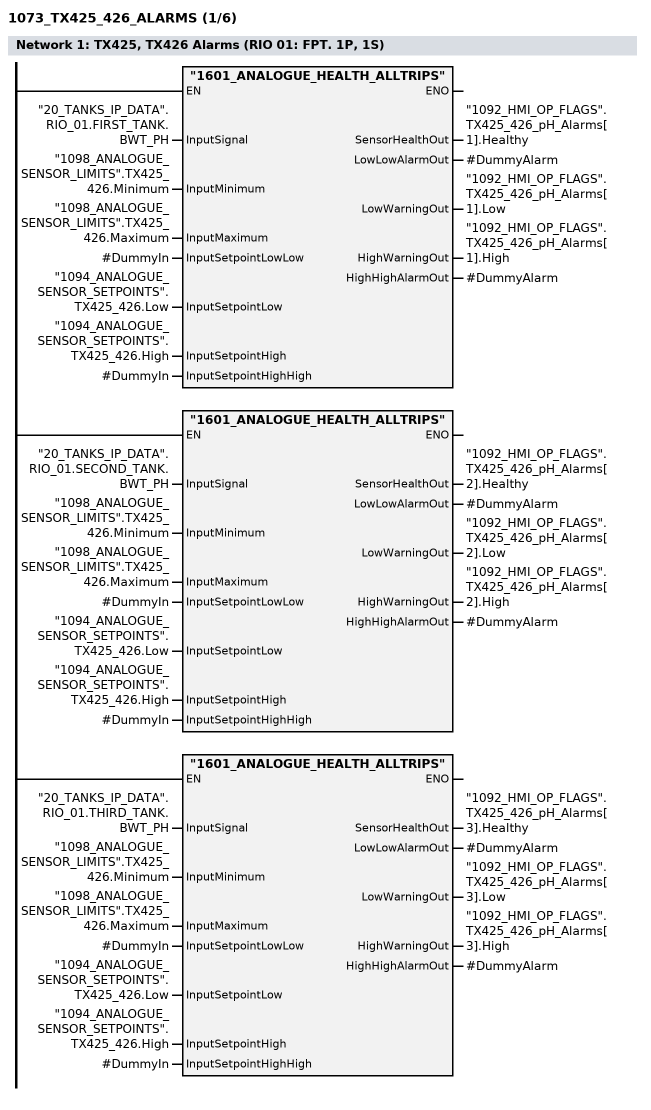
   RUNG wire#powerrail
      "1601_ANALOGUE_HEALTH_ALLTRIPS"(InputSignal := "20_TANKS_IP_DATA".RIO_01.FIRST_TANK.BWT_PH, InputMinimum := "1098_ANALOGUE_SENSOR_LIMITS".TX425_426.Minimum, InputMaximum := "1098_ANALOGUE_SENSOR_LIMITS".TX425_426.Maximum, InputSetpointLowLow := #DummyIn, InputSetpointLow := "1094_ANALOGUE_SENSOR_SETPOINTS".TX425_426.Low, InputSetpointHigh := "1094_ANALOGUE_SENSOR_SETPOINTS".TX425_426.High, InputSetpointHighHigh := #DummyIn, SensorHealthOut => "1092_HMI_OP_FLAGS".TX425_426_pH_Alarms[1].Healthy, LowLowAlarmOut => #DummyAlarm, LowWarningOut => "1092_HMI_OP_FLAGS".TX425_426_pH_Alarms[1].Low, HighWarningOut => "1092_HMI_OP_FLAGS".TX425_426_pH_Alarms[1].High, HighHighAlarmOut => #DummyAlarm)
   END_RUNG
   RUNG wire#powerrail
      "1601_ANALOGUE_HEALTH_ALLTRIPS"(InputSignal := "20_TANKS_IP_DATA".RIO_01.SECOND_TANK.BWT_PH, InputMinimum := "1098_ANALOGUE_SENSOR_LIMITS".TX425_426.Minimum, InputMaximum := "1098_ANALOGUE_SENSOR_LIMITS".TX425_426.Maximum, InputSetpointLowLow := #DummyIn, InputSetpointLow := "1094_ANALOGUE_SENSOR_SETPOINTS".TX425_426.Low, InputSetpointHigh := "1094_ANALOGUE_SENSOR_SETPOINTS".TX425_426.High, InputSetpointHighHigh := #DummyIn, SensorHealthOut => "1092_HMI_OP_FLAGS".TX425_426_pH_Alarms[2].Healthy, LowLowAlarmOut => #DummyAlarm, LowWarningOut => "1092_HMI_OP_FLAGS".TX425_426_pH_Alarms[2].Low, HighWarningOut => "1092_HMI_OP_FLAGS".TX425_426_pH_Alarms[2].High, HighHighAlarmOut => #DummyAlarm)
   END_RUNG
   RUNG wire#powerrail
      "1601_ANALOGUE_HEALTH_ALLTRIPS"(InputSignal := "20_TANKS_IP_DATA".RIO_01.THIRD_TANK.BWT_PH, InputMinimum := "1098_ANALOGUE_SENSOR_LIMITS".TX425_426.Minimum, InputMaximum := "1098_ANALOGUE_SENSOR_LIMITS".TX425_426.Maximum, InputSetpointLowLow := #DummyIn, InputSetpointLow := "1094_ANALOGUE_SENSOR_SETPOINTS".TX425_426.Low, InputSetpointHigh := "1094_ANALOGUE_SENSOR_SETPOINTS".TX425_426.High, InputSetpointHighHigh := #DummyIn, SensorHealthOut => "1092_HMI_OP_FLAGS".TX425_426_pH_Alarms[3].Healthy, LowLowAlarmOut => #DummyAlarm, LowWarningOut => "1092_HMI_OP_FLAGS".TX425_426_pH_Alarms[3].Low, HighWarningOut => "1092_HMI_OP_FLAGS".TX425_426_pH_Alarms[3].High, HighHighAlarmOut => #DummyAlarm)
   END_RUNG
   // the same network as SCL:
   "1601_ANALOGUE_HEALTH_ALLTRIPS"(InputSignal := "20_TANKS_IP_DATA".RIO_01.FIRST_TANK.BWT_PH,
                           InputMinimum := "1098_ANALOGUE_SENSOR_LIMITS".TX425_426.Minimum,
                           InputMaximum := "1098_ANALOGUE_SENSOR_LIMITS".TX425_426.Maximum,
                           InputSetpointLowLow := #DummyIn,
                           InputSetpointLow := "1094_ANALOGUE_SENSOR_SETPOINTS".TX425_426.Low,
                           InputSetpointHigh := "1094_ANALOGUE_SENSOR_SETPOINTS".TX425_426.High,
                           InputSetpointHighHigh := #DummyIn,
                           SensorHealthOut => "1092_HMI_OP_FLAGS".TX425_426_pH_Alarms[1].Healthy,
                           LowLowAlarmOut => #DummyAlarm,
                           LowWarningOut => "1092_HMI_OP_FLAGS".TX425_426_pH_Alarms[1].Low,
                           HighWarningOut => "1092_HMI_OP_FLAGS".TX425_426_pH_Alarms[1].High,
                           HighHighAlarmOut => #DummyAlarm);
   "1601_ANALOGUE_HEALTH_ALLTRIPS"(InputSignal := "20_TANKS_IP_DATA".RIO_01.SECOND_TANK.BWT_PH,
                           InputMinimum := "1098_ANALOGUE_SENSOR_LIMITS".TX425_426.Minimum,
                           InputMaximum := "1098_ANALOGUE_SENSOR_LIMITS".TX425_426.Maximum,
                           InputSetpointLowLow := #DummyIn,
                           InputSetpointLow := "1094_ANALOGUE_SENSOR_SETPOINTS".TX425_426.Low,
                           InputSetpointHigh := "1094_ANALOGUE_SENSOR_SETPOINTS".TX425_426.High,
                           InputSetpointHighHigh := #DummyIn,
                           SensorHealthOut => "1092_HMI_OP_FLAGS".TX425_426_pH_Alarms[2].Healthy,
                           LowLowAlarmOut => #DummyAlarm,
                           LowWarningOut => "1092_HMI_OP_FLAGS".TX425_426_pH_Alarms[2].Low,
                           HighWarningOut => "1092_HMI_OP_FLAGS".TX425_426_pH_Alarms[2].High,
                           HighHighAlarmOut => #DummyAlarm);
   "1601_ANALOGUE_HEALTH_ALLTRIPS"(InputSignal := "20_TANKS_IP_DATA".RIO_01.THIRD_TANK.BWT_PH,
                           InputMinimum := "1098_ANALOGUE_SENSOR_LIMITS".TX425_426.Minimum,
                           InputMaximum := "1098_ANALOGUE_SENSOR_LIMITS".TX425_426.Maximum,
                           InputSetpointLowLow := #DummyIn,
                           InputSetpointLow := "1094_ANALOGUE_SENSOR_SETPOINTS".TX425_426.Low,
                           InputSetpointHigh := "1094_ANALOGUE_SENSOR_SETPOINTS".TX425_426.High,
                           InputSetpointHighHigh := #DummyIn,
                           SensorHealthOut => "1092_HMI_OP_FLAGS".TX425_426_pH_Alarms[3].Healthy,
                           LowLowAlarmOut => #DummyAlarm,
                           LowWarningOut => "1092_HMI_OP_FLAGS".TX425_426_pH_Alarms[3].Low,
                           HighWarningOut => "1092_HMI_OP_FLAGS".TX425_426_pH_Alarms[3].High,
                           HighHighAlarmOut => #DummyAlarm);
END_REGION

REGION Network 2: TX425, TX426 Alarms (RIO 02: 2P, 2S)
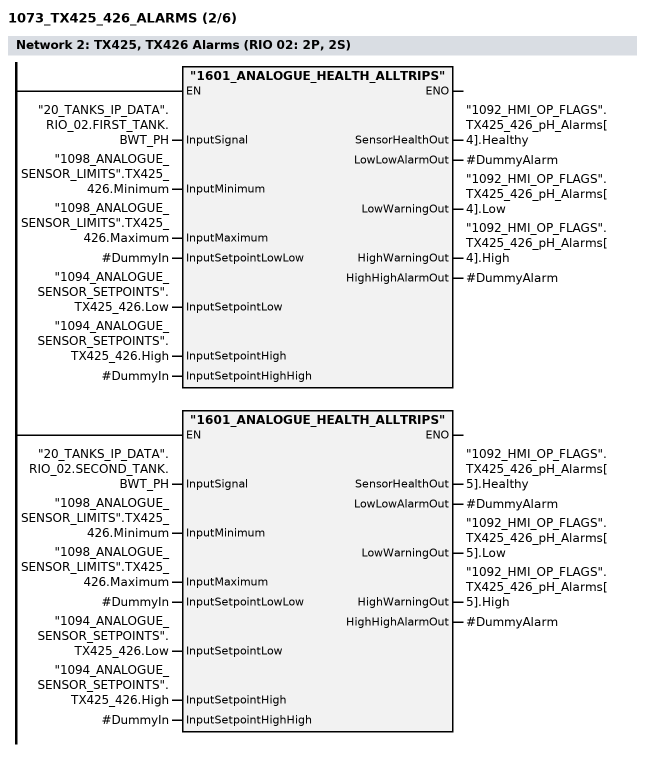
   RUNG wire#powerrail
      "1601_ANALOGUE_HEALTH_ALLTRIPS"(InputSignal := "20_TANKS_IP_DATA".RIO_02.FIRST_TANK.BWT_PH, InputMinimum := "1098_ANALOGUE_SENSOR_LIMITS".TX425_426.Minimum, InputMaximum := "1098_ANALOGUE_SENSOR_LIMITS".TX425_426.Maximum, InputSetpointLowLow := #DummyIn, InputSetpointLow := "1094_ANALOGUE_SENSOR_SETPOINTS".TX425_426.Low, InputSetpointHigh := "1094_ANALOGUE_SENSOR_SETPOINTS".TX425_426.High, InputSetpointHighHigh := #DummyIn, SensorHealthOut => "1092_HMI_OP_FLAGS".TX425_426_pH_Alarms[4].Healthy, LowLowAlarmOut => #DummyAlarm, LowWarningOut => "1092_HMI_OP_FLAGS".TX425_426_pH_Alarms[4].Low, HighWarningOut => "1092_HMI_OP_FLAGS".TX425_426_pH_Alarms[4].High, HighHighAlarmOut => #DummyAlarm)
   END_RUNG
   RUNG wire#powerrail
      "1601_ANALOGUE_HEALTH_ALLTRIPS"(InputSignal := "20_TANKS_IP_DATA".RIO_02.SECOND_TANK.BWT_PH, InputMinimum := "1098_ANALOGUE_SENSOR_LIMITS".TX425_426.Minimum, InputMaximum := "1098_ANALOGUE_SENSOR_LIMITS".TX425_426.Maximum, InputSetpointLowLow := #DummyIn, InputSetpointLow := "1094_ANALOGUE_SENSOR_SETPOINTS".TX425_426.Low, InputSetpointHigh := "1094_ANALOGUE_SENSOR_SETPOINTS".TX425_426.High, InputSetpointHighHigh := #DummyIn, SensorHealthOut => "1092_HMI_OP_FLAGS".TX425_426_pH_Alarms[5].Healthy, LowLowAlarmOut => #DummyAlarm, LowWarningOut => "1092_HMI_OP_FLAGS".TX425_426_pH_Alarms[5].Low, HighWarningOut => "1092_HMI_OP_FLAGS".TX425_426_pH_Alarms[5].High, HighHighAlarmOut => #DummyAlarm)
   END_RUNG
   // the same network as SCL:
   "1601_ANALOGUE_HEALTH_ALLTRIPS"(InputSignal := "20_TANKS_IP_DATA".RIO_02.FIRST_TANK.BWT_PH,
                           InputMinimum := "1098_ANALOGUE_SENSOR_LIMITS".TX425_426.Minimum,
                           InputMaximum := "1098_ANALOGUE_SENSOR_LIMITS".TX425_426.Maximum,
                           InputSetpointLowLow := #DummyIn,
                           InputSetpointLow := "1094_ANALOGUE_SENSOR_SETPOINTS".TX425_426.Low,
                           InputSetpointHigh := "1094_ANALOGUE_SENSOR_SETPOINTS".TX425_426.High,
                           InputSetpointHighHigh := #DummyIn,
                           SensorHealthOut => "1092_HMI_OP_FLAGS".TX425_426_pH_Alarms[4].Healthy,
                           LowLowAlarmOut => #DummyAlarm,
                           LowWarningOut => "1092_HMI_OP_FLAGS".TX425_426_pH_Alarms[4].Low,
                           HighWarningOut => "1092_HMI_OP_FLAGS".TX425_426_pH_Alarms[4].High,
                           HighHighAlarmOut => #DummyAlarm);
   "1601_ANALOGUE_HEALTH_ALLTRIPS"(InputSignal := "20_TANKS_IP_DATA".RIO_02.SECOND_TANK.BWT_PH,
                           InputMinimum := "1098_ANALOGUE_SENSOR_LIMITS".TX425_426.Minimum,
                           InputMaximum := "1098_ANALOGUE_SENSOR_LIMITS".TX425_426.Maximum,
                           InputSetpointLowLow := #DummyIn,
                           InputSetpointLow := "1094_ANALOGUE_SENSOR_SETPOINTS".TX425_426.Low,
                           InputSetpointHigh := "1094_ANALOGUE_SENSOR_SETPOINTS".TX425_426.High,
                           InputSetpointHighHigh := #DummyIn,
                           SensorHealthOut => "1092_HMI_OP_FLAGS".TX425_426_pH_Alarms[5].Healthy,
                           LowLowAlarmOut => #DummyAlarm,
                           LowWarningOut => "1092_HMI_OP_FLAGS".TX425_426_pH_Alarms[5].Low,
                           HighWarningOut => "1092_HMI_OP_FLAGS".TX425_426_pH_Alarms[5].High,
                           HighHighAlarmOut => #DummyAlarm);
END_REGION

REGION Network 3: TX425, TX426 Alarms (RIO 03: 3P, 3S)
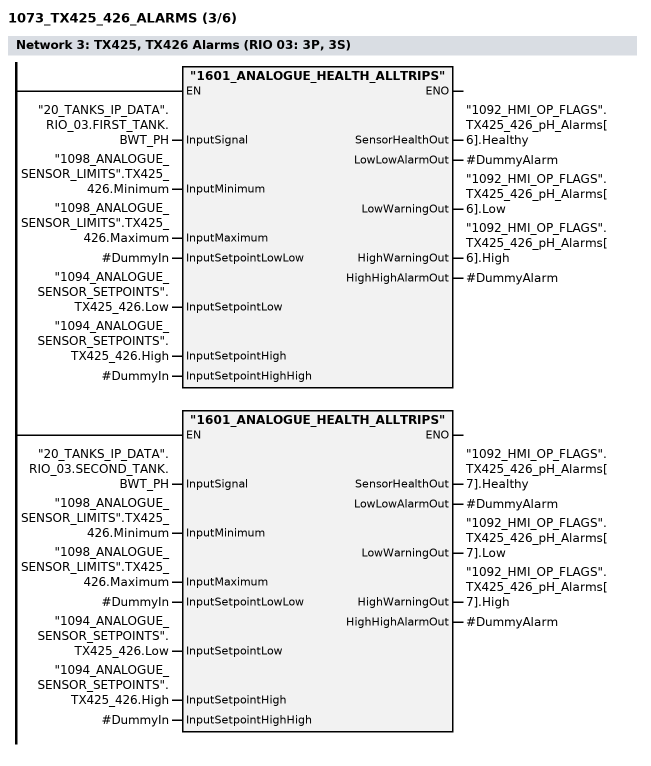
   RUNG wire#powerrail
      "1601_ANALOGUE_HEALTH_ALLTRIPS"(InputSignal := "20_TANKS_IP_DATA".RIO_03.FIRST_TANK.BWT_PH, InputMinimum := "1098_ANALOGUE_SENSOR_LIMITS".TX425_426.Minimum, InputMaximum := "1098_ANALOGUE_SENSOR_LIMITS".TX425_426.Maximum, InputSetpointLowLow := #DummyIn, InputSetpointLow := "1094_ANALOGUE_SENSOR_SETPOINTS".TX425_426.Low, InputSetpointHigh := "1094_ANALOGUE_SENSOR_SETPOINTS".TX425_426.High, InputSetpointHighHigh := #DummyIn, SensorHealthOut => "1092_HMI_OP_FLAGS".TX425_426_pH_Alarms[6].Healthy, LowLowAlarmOut => #DummyAlarm, LowWarningOut => "1092_HMI_OP_FLAGS".TX425_426_pH_Alarms[6].Low, HighWarningOut => "1092_HMI_OP_FLAGS".TX425_426_pH_Alarms[6].High, HighHighAlarmOut => #DummyAlarm)
   END_RUNG
   RUNG wire#powerrail
      "1601_ANALOGUE_HEALTH_ALLTRIPS"(InputSignal := "20_TANKS_IP_DATA".RIO_03.SECOND_TANK.BWT_PH, InputMinimum := "1098_ANALOGUE_SENSOR_LIMITS".TX425_426.Minimum, InputMaximum := "1098_ANALOGUE_SENSOR_LIMITS".TX425_426.Maximum, InputSetpointLowLow := #DummyIn, InputSetpointLow := "1094_ANALOGUE_SENSOR_SETPOINTS".TX425_426.Low, InputSetpointHigh := "1094_ANALOGUE_SENSOR_SETPOINTS".TX425_426.High, InputSetpointHighHigh := #DummyIn, SensorHealthOut => "1092_HMI_OP_FLAGS".TX425_426_pH_Alarms[7].Healthy, LowLowAlarmOut => #DummyAlarm, LowWarningOut => "1092_HMI_OP_FLAGS".TX425_426_pH_Alarms[7].Low, HighWarningOut => "1092_HMI_OP_FLAGS".TX425_426_pH_Alarms[7].High, HighHighAlarmOut => #DummyAlarm)
   END_RUNG
   // the same network as SCL:
   "1601_ANALOGUE_HEALTH_ALLTRIPS"(InputSignal := "20_TANKS_IP_DATA".RIO_03.FIRST_TANK.BWT_PH,
                           InputMinimum := "1098_ANALOGUE_SENSOR_LIMITS".TX425_426.Minimum,
                           InputMaximum := "1098_ANALOGUE_SENSOR_LIMITS".TX425_426.Maximum,
                           InputSetpointLowLow := #DummyIn,
                           InputSetpointLow := "1094_ANALOGUE_SENSOR_SETPOINTS".TX425_426.Low,
                           InputSetpointHigh := "1094_ANALOGUE_SENSOR_SETPOINTS".TX425_426.High,
                           InputSetpointHighHigh := #DummyIn,
                           SensorHealthOut => "1092_HMI_OP_FLAGS".TX425_426_pH_Alarms[6].Healthy,
                           LowLowAlarmOut => #DummyAlarm,
                           LowWarningOut => "1092_HMI_OP_FLAGS".TX425_426_pH_Alarms[6].Low,
                           HighWarningOut => "1092_HMI_OP_FLAGS".TX425_426_pH_Alarms[6].High,
                           HighHighAlarmOut => #DummyAlarm);
   "1601_ANALOGUE_HEALTH_ALLTRIPS"(InputSignal := "20_TANKS_IP_DATA".RIO_03.SECOND_TANK.BWT_PH,
                           InputMinimum := "1098_ANALOGUE_SENSOR_LIMITS".TX425_426.Minimum,
                           InputMaximum := "1098_ANALOGUE_SENSOR_LIMITS".TX425_426.Maximum,
                           InputSetpointLowLow := #DummyIn,
                           InputSetpointLow := "1094_ANALOGUE_SENSOR_SETPOINTS".TX425_426.Low,
                           InputSetpointHigh := "1094_ANALOGUE_SENSOR_SETPOINTS".TX425_426.High,
                           InputSetpointHighHigh := #DummyIn,
                           SensorHealthOut => "1092_HMI_OP_FLAGS".TX425_426_pH_Alarms[7].Healthy,
                           LowLowAlarmOut => #DummyAlarm,
                           LowWarningOut => "1092_HMI_OP_FLAGS".TX425_426_pH_Alarms[7].Low,
                           HighWarningOut => "1092_HMI_OP_FLAGS".TX425_426_pH_Alarms[7].High,
                           HighHighAlarmOut => #DummyAlarm);
END_REGION

REGION Network 4: TX425, TX426 Alarms (RIO 04: 4P, 4S)
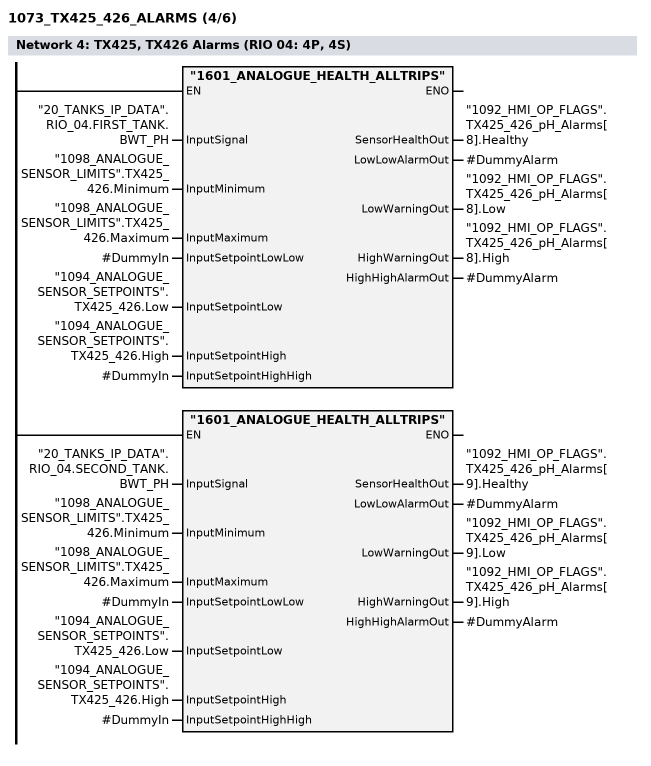
   RUNG wire#powerrail
      "1601_ANALOGUE_HEALTH_ALLTRIPS"(InputSignal := "20_TANKS_IP_DATA".RIO_04.FIRST_TANK.BWT_PH, InputMinimum := "1098_ANALOGUE_SENSOR_LIMITS".TX425_426.Minimum, InputMaximum := "1098_ANALOGUE_SENSOR_LIMITS".TX425_426.Maximum, InputSetpointLowLow := #DummyIn, InputSetpointLow := "1094_ANALOGUE_SENSOR_SETPOINTS".TX425_426.Low, InputSetpointHigh := "1094_ANALOGUE_SENSOR_SETPOINTS".TX425_426.High, InputSetpointHighHigh := #DummyIn, SensorHealthOut => "1092_HMI_OP_FLAGS".TX425_426_pH_Alarms[8].Healthy, LowLowAlarmOut => #DummyAlarm, LowWarningOut => "1092_HMI_OP_FLAGS".TX425_426_pH_Alarms[8].Low, HighWarningOut => "1092_HMI_OP_FLAGS".TX425_426_pH_Alarms[8].High, HighHighAlarmOut => #DummyAlarm)
   END_RUNG
   RUNG wire#powerrail
      "1601_ANALOGUE_HEALTH_ALLTRIPS"(InputSignal := "20_TANKS_IP_DATA".RIO_04.SECOND_TANK.BWT_PH, InputMinimum := "1098_ANALOGUE_SENSOR_LIMITS".TX425_426.Minimum, InputMaximum := "1098_ANALOGUE_SENSOR_LIMITS".TX425_426.Maximum, InputSetpointLowLow := #DummyIn, InputSetpointLow := "1094_ANALOGUE_SENSOR_SETPOINTS".TX425_426.Low, InputSetpointHigh := "1094_ANALOGUE_SENSOR_SETPOINTS".TX425_426.High, InputSetpointHighHigh := #DummyIn, SensorHealthOut => "1092_HMI_OP_FLAGS".TX425_426_pH_Alarms[9].Healthy, LowLowAlarmOut => #DummyAlarm, LowWarningOut => "1092_HMI_OP_FLAGS".TX425_426_pH_Alarms[9].Low, HighWarningOut => "1092_HMI_OP_FLAGS".TX425_426_pH_Alarms[9].High, HighHighAlarmOut => #DummyAlarm)
   END_RUNG
   // the same network as SCL:
   "1601_ANALOGUE_HEALTH_ALLTRIPS"(InputSignal := "20_TANKS_IP_DATA".RIO_04.FIRST_TANK.BWT_PH,
                           InputMinimum := "1098_ANALOGUE_SENSOR_LIMITS".TX425_426.Minimum,
                           InputMaximum := "1098_ANALOGUE_SENSOR_LIMITS".TX425_426.Maximum,
                           InputSetpointLowLow := #DummyIn,
                           InputSetpointLow := "1094_ANALOGUE_SENSOR_SETPOINTS".TX425_426.Low,
                           InputSetpointHigh := "1094_ANALOGUE_SENSOR_SETPOINTS".TX425_426.High,
                           InputSetpointHighHigh := #DummyIn,
                           SensorHealthOut => "1092_HMI_OP_FLAGS".TX425_426_pH_Alarms[8].Healthy,
                           LowLowAlarmOut => #DummyAlarm,
                           LowWarningOut => "1092_HMI_OP_FLAGS".TX425_426_pH_Alarms[8].Low,
                           HighWarningOut => "1092_HMI_OP_FLAGS".TX425_426_pH_Alarms[8].High,
                           HighHighAlarmOut => #DummyAlarm);
   "1601_ANALOGUE_HEALTH_ALLTRIPS"(InputSignal := "20_TANKS_IP_DATA".RIO_04.SECOND_TANK.BWT_PH,
                           InputMinimum := "1098_ANALOGUE_SENSOR_LIMITS".TX425_426.Minimum,
                           InputMaximum := "1098_ANALOGUE_SENSOR_LIMITS".TX425_426.Maximum,
                           InputSetpointLowLow := #DummyIn,
                           InputSetpointLow := "1094_ANALOGUE_SENSOR_SETPOINTS".TX425_426.Low,
                           InputSetpointHigh := "1094_ANALOGUE_SENSOR_SETPOINTS".TX425_426.High,
                           InputSetpointHighHigh := #DummyIn,
                           SensorHealthOut => "1092_HMI_OP_FLAGS".TX425_426_pH_Alarms[9].Healthy,
                           LowLowAlarmOut => #DummyAlarm,
                           LowWarningOut => "1092_HMI_OP_FLAGS".TX425_426_pH_Alarms[9].Low,
                           HighWarningOut => "1092_HMI_OP_FLAGS".TX425_426_pH_Alarms[9].High,
                           HighHighAlarmOut => #DummyAlarm);
END_REGION

REGION Network 5: TX425, TX426 Alarms (RIO 05: 5P, 5S)
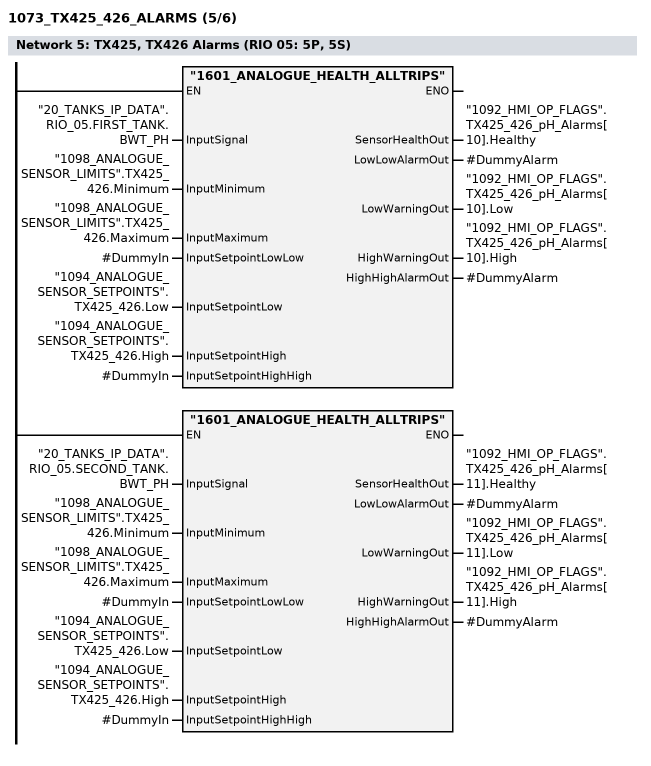
   RUNG wire#powerrail
      "1601_ANALOGUE_HEALTH_ALLTRIPS"(InputSignal := "20_TANKS_IP_DATA".RIO_05.FIRST_TANK.BWT_PH, InputMinimum := "1098_ANALOGUE_SENSOR_LIMITS".TX425_426.Minimum, InputMaximum := "1098_ANALOGUE_SENSOR_LIMITS".TX425_426.Maximum, InputSetpointLowLow := #DummyIn, InputSetpointLow := "1094_ANALOGUE_SENSOR_SETPOINTS".TX425_426.Low, InputSetpointHigh := "1094_ANALOGUE_SENSOR_SETPOINTS".TX425_426.High, InputSetpointHighHigh := #DummyIn, SensorHealthOut => "1092_HMI_OP_FLAGS".TX425_426_pH_Alarms[10].Healthy, LowLowAlarmOut => #DummyAlarm, LowWarningOut => "1092_HMI_OP_FLAGS".TX425_426_pH_Alarms[10].Low, HighWarningOut => "1092_HMI_OP_FLAGS".TX425_426_pH_Alarms[10].High, HighHighAlarmOut => #DummyAlarm)
   END_RUNG
   RUNG wire#powerrail
      "1601_ANALOGUE_HEALTH_ALLTRIPS"(InputSignal := "20_TANKS_IP_DATA".RIO_05.SECOND_TANK.BWT_PH, InputMinimum := "1098_ANALOGUE_SENSOR_LIMITS".TX425_426.Minimum, InputMaximum := "1098_ANALOGUE_SENSOR_LIMITS".TX425_426.Maximum, InputSetpointLowLow := #DummyIn, InputSetpointLow := "1094_ANALOGUE_SENSOR_SETPOINTS".TX425_426.Low, InputSetpointHigh := "1094_ANALOGUE_SENSOR_SETPOINTS".TX425_426.High, InputSetpointHighHigh := #DummyIn, SensorHealthOut => "1092_HMI_OP_FLAGS".TX425_426_pH_Alarms[11].Healthy, LowLowAlarmOut => #DummyAlarm, LowWarningOut => "1092_HMI_OP_FLAGS".TX425_426_pH_Alarms[11].Low, HighWarningOut => "1092_HMI_OP_FLAGS".TX425_426_pH_Alarms[11].High, HighHighAlarmOut => #DummyAlarm)
   END_RUNG
   // the same network as SCL:
   "1601_ANALOGUE_HEALTH_ALLTRIPS"(InputSignal := "20_TANKS_IP_DATA".RIO_05.FIRST_TANK.BWT_PH,
                           InputMinimum := "1098_ANALOGUE_SENSOR_LIMITS".TX425_426.Minimum,
                           InputMaximum := "1098_ANALOGUE_SENSOR_LIMITS".TX425_426.Maximum,
                           InputSetpointLowLow := #DummyIn,
                           InputSetpointLow := "1094_ANALOGUE_SENSOR_SETPOINTS".TX425_426.Low,
                           InputSetpointHigh := "1094_ANALOGUE_SENSOR_SETPOINTS".TX425_426.High,
                           InputSetpointHighHigh := #DummyIn,
                           SensorHealthOut => "1092_HMI_OP_FLAGS".TX425_426_pH_Alarms[10].Healthy,
                           LowLowAlarmOut => #DummyAlarm,
                           LowWarningOut => "1092_HMI_OP_FLAGS".TX425_426_pH_Alarms[10].Low,
                           HighWarningOut => "1092_HMI_OP_FLAGS".TX425_426_pH_Alarms[10].High,
                           HighHighAlarmOut => #DummyAlarm);
   "1601_ANALOGUE_HEALTH_ALLTRIPS"(InputSignal := "20_TANKS_IP_DATA".RIO_05.SECOND_TANK.BWT_PH,
                           InputMinimum := "1098_ANALOGUE_SENSOR_LIMITS".TX425_426.Minimum,
                           InputMaximum := "1098_ANALOGUE_SENSOR_LIMITS".TX425_426.Maximum,
                           InputSetpointLowLow := #DummyIn,
                           InputSetpointLow := "1094_ANALOGUE_SENSOR_SETPOINTS".TX425_426.Low,
                           InputSetpointHigh := "1094_ANALOGUE_SENSOR_SETPOINTS".TX425_426.High,
                           InputSetpointHighHigh := #DummyIn,
                           SensorHealthOut => "1092_HMI_OP_FLAGS".TX425_426_pH_Alarms[11].Healthy,
                           LowLowAlarmOut => #DummyAlarm,
                           LowWarningOut => "1092_HMI_OP_FLAGS".TX425_426_pH_Alarms[11].Low,
                           HighWarningOut => "1092_HMI_OP_FLAGS".TX425_426_pH_Alarms[11].High,
                           HighHighAlarmOut => #DummyAlarm);
END_REGION

REGION Network 6: TX425, TX426 Alarms (RIO 06: 6P, 6S)
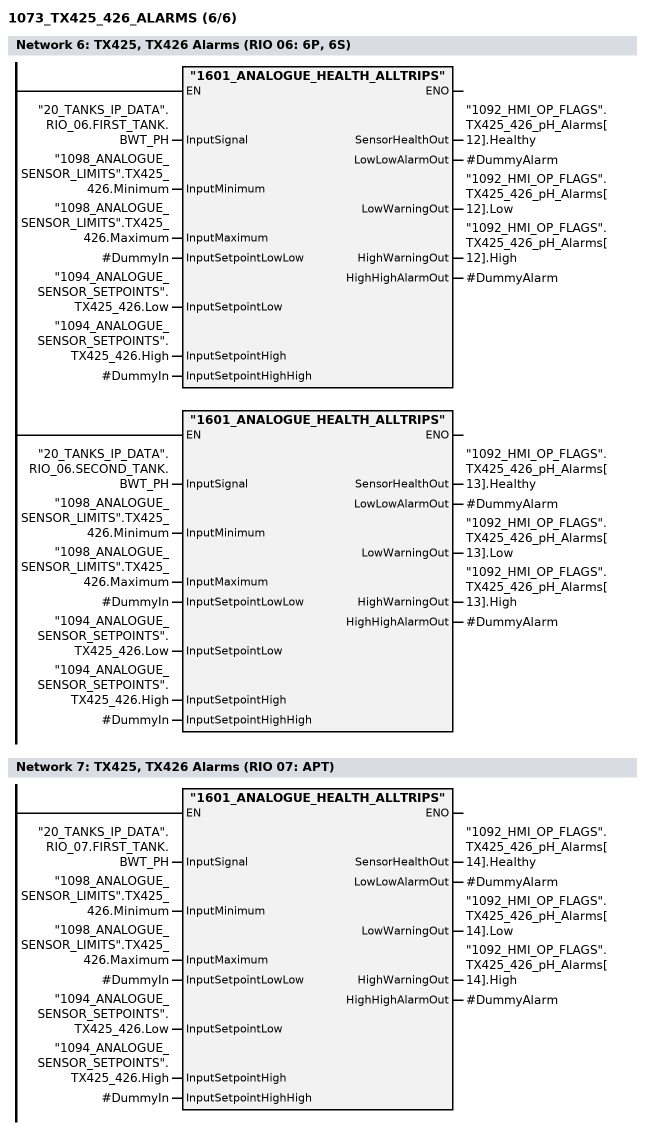
   RUNG wire#powerrail
      "1601_ANALOGUE_HEALTH_ALLTRIPS"(InputSignal := "20_TANKS_IP_DATA".RIO_06.FIRST_TANK.BWT_PH, InputMinimum := "1098_ANALOGUE_SENSOR_LIMITS".TX425_426.Minimum, InputMaximum := "1098_ANALOGUE_SENSOR_LIMITS".TX425_426.Maximum, InputSetpointLowLow := #DummyIn, InputSetpointLow := "1094_ANALOGUE_SENSOR_SETPOINTS".TX425_426.Low, InputSetpointHigh := "1094_ANALOGUE_SENSOR_SETPOINTS".TX425_426.High, InputSetpointHighHigh := #DummyIn, SensorHealthOut => "1092_HMI_OP_FLAGS".TX425_426_pH_Alarms[12].Healthy, LowLowAlarmOut => #DummyAlarm, LowWarningOut => "1092_HMI_OP_FLAGS".TX425_426_pH_Alarms[12].Low, HighWarningOut => "1092_HMI_OP_FLAGS".TX425_426_pH_Alarms[12].High, HighHighAlarmOut => #DummyAlarm)
   END_RUNG
   RUNG wire#powerrail
      "1601_ANALOGUE_HEALTH_ALLTRIPS"(InputSignal := "20_TANKS_IP_DATA".RIO_06.SECOND_TANK.BWT_PH, InputMinimum := "1098_ANALOGUE_SENSOR_LIMITS".TX425_426.Minimum, InputMaximum := "1098_ANALOGUE_SENSOR_LIMITS".TX425_426.Maximum, InputSetpointLowLow := #DummyIn, InputSetpointLow := "1094_ANALOGUE_SENSOR_SETPOINTS".TX425_426.Low, InputSetpointHigh := "1094_ANALOGUE_SENSOR_SETPOINTS".TX425_426.High, InputSetpointHighHigh := #DummyIn, SensorHealthOut => "1092_HMI_OP_FLAGS".TX425_426_pH_Alarms[13].Healthy, LowLowAlarmOut => #DummyAlarm, LowWarningOut => "1092_HMI_OP_FLAGS".TX425_426_pH_Alarms[13].Low, HighWarningOut => "1092_HMI_OP_FLAGS".TX425_426_pH_Alarms[13].High, HighHighAlarmOut => #DummyAlarm)
   END_RUNG
   // the same network as SCL:
   "1601_ANALOGUE_HEALTH_ALLTRIPS"(InputSignal := "20_TANKS_IP_DATA".RIO_06.FIRST_TANK.BWT_PH,
                           InputMinimum := "1098_ANALOGUE_SENSOR_LIMITS".TX425_426.Minimum,
                           InputMaximum := "1098_ANALOGUE_SENSOR_LIMITS".TX425_426.Maximum,
                           InputSetpointLowLow := #DummyIn,
                           InputSetpointLow := "1094_ANALOGUE_SENSOR_SETPOINTS".TX425_426.Low,
                           InputSetpointHigh := "1094_ANALOGUE_SENSOR_SETPOINTS".TX425_426.High,
                           InputSetpointHighHigh := #DummyIn,
                           SensorHealthOut => "1092_HMI_OP_FLAGS".TX425_426_pH_Alarms[12].Healthy,
                           LowLowAlarmOut => #DummyAlarm,
                           LowWarningOut => "1092_HMI_OP_FLAGS".TX425_426_pH_Alarms[12].Low,
                           HighWarningOut => "1092_HMI_OP_FLAGS".TX425_426_pH_Alarms[12].High,
                           HighHighAlarmOut => #DummyAlarm);
   "1601_ANALOGUE_HEALTH_ALLTRIPS"(InputSignal := "20_TANKS_IP_DATA".RIO_06.SECOND_TANK.BWT_PH,
                           InputMinimum := "1098_ANALOGUE_SENSOR_LIMITS".TX425_426.Minimum,
                           InputMaximum := "1098_ANALOGUE_SENSOR_LIMITS".TX425_426.Maximum,
                           InputSetpointLowLow := #DummyIn,
                           InputSetpointLow := "1094_ANALOGUE_SENSOR_SETPOINTS".TX425_426.Low,
                           InputSetpointHigh := "1094_ANALOGUE_SENSOR_SETPOINTS".TX425_426.High,
                           InputSetpointHighHigh := #DummyIn,
                           SensorHealthOut => "1092_HMI_OP_FLAGS".TX425_426_pH_Alarms[13].Healthy,
                           LowLowAlarmOut => #DummyAlarm,
                           LowWarningOut => "1092_HMI_OP_FLAGS".TX425_426_pH_Alarms[13].Low,
                           HighWarningOut => "1092_HMI_OP_FLAGS".TX425_426_pH_Alarms[13].High,
                           HighHighAlarmOut => #DummyAlarm);
END_REGION

REGION Network 7: TX425, TX426 Alarms (RIO 07: APT)
   RUNG wire#powerrail
      "1601_ANALOGUE_HEALTH_ALLTRIPS"(InputSignal := "20_TANKS_IP_DATA".RIO_07.FIRST_TANK.BWT_PH, InputMinimum := "1098_ANALOGUE_SENSOR_LIMITS".TX425_426.Minimum, InputMaximum := "1098_ANALOGUE_SENSOR_LIMITS".TX425_426.Maximum, InputSetpointLowLow := #DummyIn, InputSetpointLow := "1094_ANALOGUE_SENSOR_SETPOINTS".TX425_426.Low, InputSetpointHigh := "1094_ANALOGUE_SENSOR_SETPOINTS".TX425_426.High, InputSetpointHighHigh := #DummyIn, SensorHealthOut => "1092_HMI_OP_FLAGS".TX425_426_pH_Alarms[14].Healthy, LowLowAlarmOut => #DummyAlarm, LowWarningOut => "1092_HMI_OP_FLAGS".TX425_426_pH_Alarms[14].Low, HighWarningOut => "1092_HMI_OP_FLAGS".TX425_426_pH_Alarms[14].High, HighHighAlarmOut => #DummyAlarm)
   END_RUNG
   // the same network as SCL:
   "1601_ANALOGUE_HEALTH_ALLTRIPS"(InputSignal := "20_TANKS_IP_DATA".RIO_07.FIRST_TANK.BWT_PH,
                           InputMinimum := "1098_ANALOGUE_SENSOR_LIMITS".TX425_426.Minimum,
                           InputMaximum := "1098_ANALOGUE_SENSOR_LIMITS".TX425_426.Maximum,
                           InputSetpointLowLow := #DummyIn,
                           InputSetpointLow := "1094_ANALOGUE_SENSOR_SETPOINTS".TX425_426.Low,
                           InputSetpointHigh := "1094_ANALOGUE_SENSOR_SETPOINTS".TX425_426.High,
                           InputSetpointHighHigh := #DummyIn,
                           SensorHealthOut => "1092_HMI_OP_FLAGS".TX425_426_pH_Alarms[14].Healthy,
                           LowLowAlarmOut => #DummyAlarm,
                           LowWarningOut => "1092_HMI_OP_FLAGS".TX425_426_pH_Alarms[14].Low,
                           HighWarningOut => "1092_HMI_OP_FLAGS".TX425_426_pH_Alarms[14].High,
                           HighHighAlarmOut => #DummyAlarm);
END_REGION
END_FUNCTION

FUNCTION "1074_TX427_428_ALARMS" : Void   // FC1074, LAD
{ S7_Optimized_Access := 'TRUE' }
VERSION : 0.1
// Alarm wrapper function for DO level on each tank.
// DummyIn and DummyAlarm are used to manage the unused I/O in the analog health trips function as this function only uses Low and High warnings, it does not output HighHigh or LowLow alarms.
// Note: TX427 and TX428 use differing setpoints based on the system operation mode.
   VAR_TEMP
      DummyIn : Real;   // Dummy input used if alarms are Low and High only.
      DummyAlarm : Bool;   // Dummy output used if alarms are Low and High only.
      TX427_428_SP_FPT : "ANALOG_SENSOR_SETPOINTS";
      TX427_428_SP_1P : "ANALOG_SENSOR_SETPOINTS";
      TX427_428_SP_1S : "ANALOG_SENSOR_SETPOINTS";
      TX427_428_SP_2P : "ANALOG_SENSOR_SETPOINTS";
      TX427_428_SP_2S : "ANALOG_SENSOR_SETPOINTS";
      TX427_428_SP_3P : "ANALOG_SENSOR_SETPOINTS";
      TX427_428_SP_3S : "ANALOG_SENSOR_SETPOINTS";
      TX427_428_SP_4P : "ANALOG_SENSOR_SETPOINTS";
      TX427_428_SP_4S : "ANALOG_SENSOR_SETPOINTS";
      TX427_428_SP_5P : "ANALOG_SENSOR_SETPOINTS";
      TX427_428_SP_5S : "ANALOG_SENSOR_SETPOINTS";
      TX427_428_SP_6P : "ANALOG_SENSOR_SETPOINTS";
      TX427_428_SP_6S : "ANALOG_SENSOR_SETPOINTS";
      TX427_428_SP_APT : "ANALOG_SENSOR_SETPOINTS";
   END_VAR
   VAR_TEMP   // added for the SCL form of the ladder/FBD networks
      _w1 : Bool;
      _w2 : Bool;
      _w3 : Bool;
   END_VAR
BEGIN

REGION Network 1: TX427, TX428 Alarms (RIO 01: FPT. 1P, 1S)
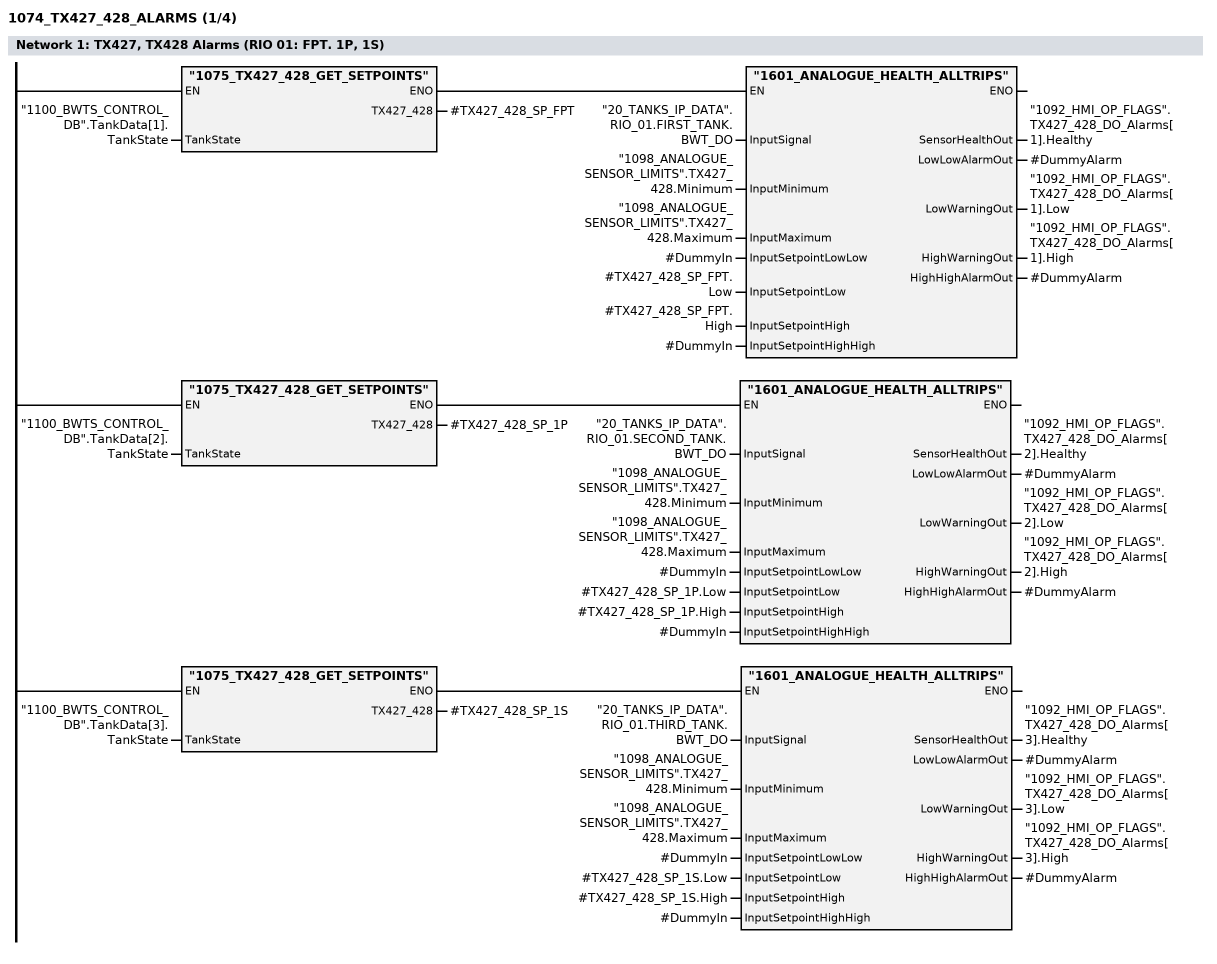
   RUNG wire#powerrail
      "1075_TX427_428_GET_SETPOINTS"(TankState := "1100_BWTS_CONTROL_DB".TankData[1].TankState, TX427_428 => #TX427_428_SP_FPT)
      "1601_ANALOGUE_HEALTH_ALLTRIPS"(InputSignal := "20_TANKS_IP_DATA".RIO_01.FIRST_TANK.BWT_DO, InputMinimum := "1098_ANALOGUE_SENSOR_LIMITS".TX427_428.Minimum, InputMaximum := "1098_ANALOGUE_SENSOR_LIMITS".TX427_428.Maximum, InputSetpointLowLow := #DummyIn, InputSetpointLow := #TX427_428_SP_FPT.Low, InputSetpointHigh := #TX427_428_SP_FPT.High, InputSetpointHighHigh := #DummyIn, SensorHealthOut => "1092_HMI_OP_FLAGS".TX427_428_DO_Alarms[1].Healthy, LowLowAlarmOut => #DummyAlarm, LowWarningOut => "1092_HMI_OP_FLAGS".TX427_428_DO_Alarms[1].Low, HighWarningOut => "1092_HMI_OP_FLAGS".TX427_428_DO_Alarms[1].High, HighHighAlarmOut => #DummyAlarm)
   END_RUNG
   RUNG wire#powerrail
      "1075_TX427_428_GET_SETPOINTS"(TankState := "1100_BWTS_CONTROL_DB".TankData[2].TankState, TX427_428 => #TX427_428_SP_1P)
      "1601_ANALOGUE_HEALTH_ALLTRIPS"(InputSignal := "20_TANKS_IP_DATA".RIO_01.SECOND_TANK.BWT_DO, InputMinimum := "1098_ANALOGUE_SENSOR_LIMITS".TX427_428.Minimum, InputMaximum := "1098_ANALOGUE_SENSOR_LIMITS".TX427_428.Maximum, InputSetpointLowLow := #DummyIn, InputSetpointLow := #TX427_428_SP_1P.Low, InputSetpointHigh := #TX427_428_SP_1P.High, InputSetpointHighHigh := #DummyIn, SensorHealthOut => "1092_HMI_OP_FLAGS".TX427_428_DO_Alarms[2].Healthy, LowLowAlarmOut => #DummyAlarm, LowWarningOut => "1092_HMI_OP_FLAGS".TX427_428_DO_Alarms[2].Low, HighWarningOut => "1092_HMI_OP_FLAGS".TX427_428_DO_Alarms[2].High, HighHighAlarmOut => #DummyAlarm)
   END_RUNG
   RUNG wire#powerrail
      "1075_TX427_428_GET_SETPOINTS"(TankState := "1100_BWTS_CONTROL_DB".TankData[3].TankState, TX427_428 => #TX427_428_SP_1S)
      "1601_ANALOGUE_HEALTH_ALLTRIPS"(InputSignal := "20_TANKS_IP_DATA".RIO_01.THIRD_TANK.BWT_DO, InputMinimum := "1098_ANALOGUE_SENSOR_LIMITS".TX427_428.Minimum, InputMaximum := "1098_ANALOGUE_SENSOR_LIMITS".TX427_428.Maximum, InputSetpointLowLow := #DummyIn, InputSetpointLow := #TX427_428_SP_1S.Low, InputSetpointHigh := #TX427_428_SP_1S.High, InputSetpointHighHigh := #DummyIn, SensorHealthOut => "1092_HMI_OP_FLAGS".TX427_428_DO_Alarms[3].Healthy, LowLowAlarmOut => #DummyAlarm, LowWarningOut => "1092_HMI_OP_FLAGS".TX427_428_DO_Alarms[3].Low, HighWarningOut => "1092_HMI_OP_FLAGS".TX427_428_DO_Alarms[3].High, HighHighAlarmOut => #DummyAlarm)
   END_RUNG
   // the same network as SCL:
   "1075_TX427_428_GET_SETPOINTS"(TankState := "1100_BWTS_CONTROL_DB".TankData[1].TankState,
                           TX427_428 => #TX427_428_SP_FPT,
                           ENO => #_w1);
   IF #_w1 THEN
       "1601_ANALOGUE_HEALTH_ALLTRIPS"(InputSignal := "20_TANKS_IP_DATA".RIO_01.FIRST_TANK.BWT_DO,
                               InputMinimum := "1098_ANALOGUE_SENSOR_LIMITS".TX427_428.Minimum,
                               InputMaximum := "1098_ANALOGUE_SENSOR_LIMITS".TX427_428.Maximum,
                               InputSetpointLowLow := #DummyIn,
                               InputSetpointLow := #TX427_428_SP_FPT.Low,
                               InputSetpointHigh := #TX427_428_SP_FPT.High,
                               InputSetpointHighHigh := #DummyIn,
                               SensorHealthOut => "1092_HMI_OP_FLAGS".TX427_428_DO_Alarms[1].Healthy,
                               LowLowAlarmOut => #DummyAlarm,
                               LowWarningOut => "1092_HMI_OP_FLAGS".TX427_428_DO_Alarms[1].Low,
                               HighWarningOut => "1092_HMI_OP_FLAGS".TX427_428_DO_Alarms[1].High,
                               HighHighAlarmOut => #DummyAlarm);
   END_IF;
   "1075_TX427_428_GET_SETPOINTS"(TankState := "1100_BWTS_CONTROL_DB".TankData[2].TankState,
                           TX427_428 => #TX427_428_SP_1P,
                           ENO => #_w2);
   IF #_w2 THEN
       "1601_ANALOGUE_HEALTH_ALLTRIPS"(InputSignal := "20_TANKS_IP_DATA".RIO_01.SECOND_TANK.BWT_DO,
                               InputMinimum := "1098_ANALOGUE_SENSOR_LIMITS".TX427_428.Minimum,
                               InputMaximum := "1098_ANALOGUE_SENSOR_LIMITS".TX427_428.Maximum,
                               InputSetpointLowLow := #DummyIn,
                               InputSetpointLow := #TX427_428_SP_1P.Low,
                               InputSetpointHigh := #TX427_428_SP_1P.High,
                               InputSetpointHighHigh := #DummyIn,
                               SensorHealthOut => "1092_HMI_OP_FLAGS".TX427_428_DO_Alarms[2].Healthy,
                               LowLowAlarmOut => #DummyAlarm,
                               LowWarningOut => "1092_HMI_OP_FLAGS".TX427_428_DO_Alarms[2].Low,
                               HighWarningOut => "1092_HMI_OP_FLAGS".TX427_428_DO_Alarms[2].High,
                               HighHighAlarmOut => #DummyAlarm);
   END_IF;
   "1075_TX427_428_GET_SETPOINTS"(TankState := "1100_BWTS_CONTROL_DB".TankData[3].TankState,
                           TX427_428 => #TX427_428_SP_1S,
                           ENO => #_w3);
   IF #_w3 THEN
       "1601_ANALOGUE_HEALTH_ALLTRIPS"(InputSignal := "20_TANKS_IP_DATA".RIO_01.THIRD_TANK.BWT_DO,
                               InputMinimum := "1098_ANALOGUE_SENSOR_LIMITS".TX427_428.Minimum,
                               InputMaximum := "1098_ANALOGUE_SENSOR_LIMITS".TX427_428.Maximum,
                               InputSetpointLowLow := #DummyIn,
                               InputSetpointLow := #TX427_428_SP_1S.Low,
                               InputSetpointHigh := #TX427_428_SP_1S.High,
                               InputSetpointHighHigh := #DummyIn,
                               SensorHealthOut => "1092_HMI_OP_FLAGS".TX427_428_DO_Alarms[3].Healthy,
                               LowLowAlarmOut => #DummyAlarm,
                               LowWarningOut => "1092_HMI_OP_FLAGS".TX427_428_DO_Alarms[3].Low,
                               HighWarningOut => "1092_HMI_OP_FLAGS".TX427_428_DO_Alarms[3].High,
                               HighHighAlarmOut => #DummyAlarm);
   END_IF;
END_REGION

REGION Network 2: TX427, TX428 Alarms (RIO 02: 2P, 2S)